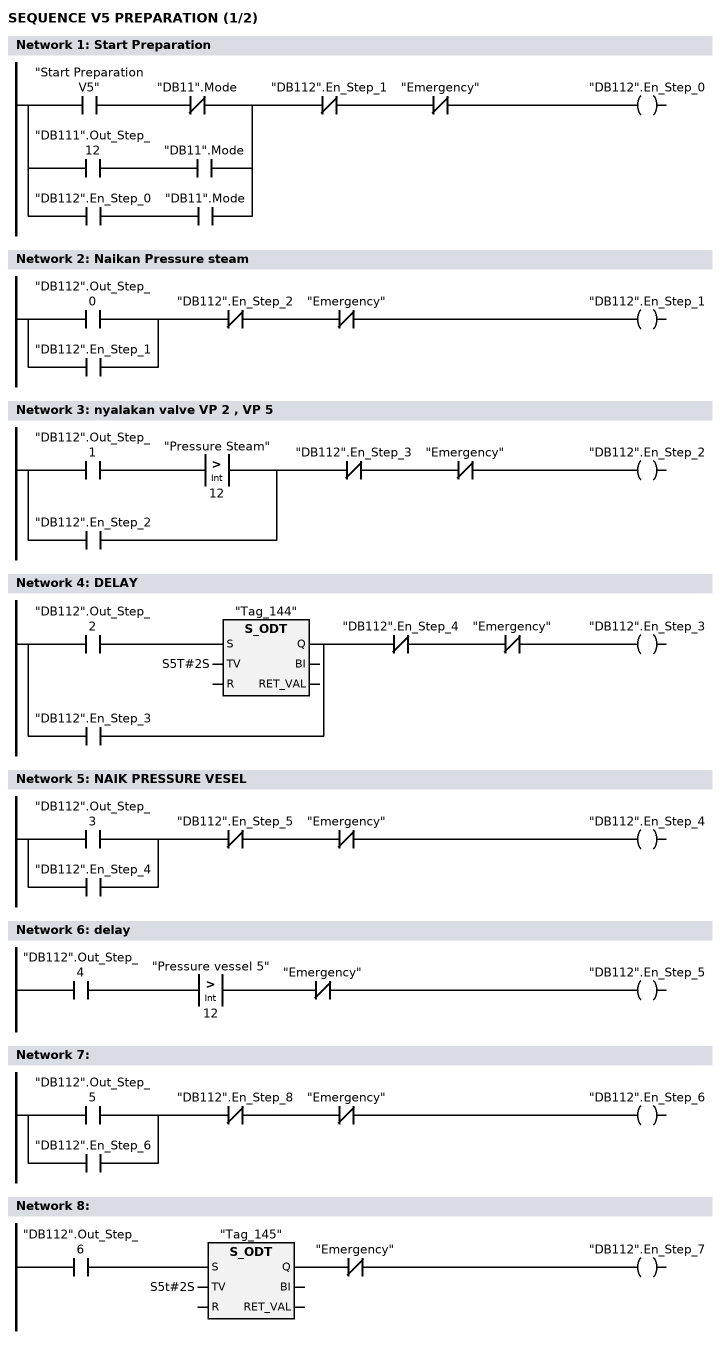
   RUNG wire#powerrail
      Contact( "Start Preparation V5" )
      I_Contact( "DB11".Mode )
      wire#w1
      I_Contact( "DB112".En_Step_1 )
      I_Contact( "Emergency" )
      Coil( "DB112".En_Step_0 )
   END_RUNG
   RUNG wire#powerrail
      Contact( "DB111".Out_Step_12 )
      Contact( "DB11".Mode )
   END_RUNG wire#w1
   RUNG wire#powerrail
      Contact( "DB112".En_Step_0 )
      Contact( "DB11".Mode )
   END_RUNG wire#w1
   // the same network as SCL:
   "DB112".En_Step_0 := (("Start Preparation V5" AND NOT "DB11".Mode) OR ("DB111".Out_Step_12 AND "DB11".Mode) OR ("DB112".En_Step_0 AND "DB11".Mode)) AND NOT "DB112".En_Step_1 AND NOT "Emergency";
END_REGION

REGION Network 2: Naikan Pressure steam
   RUNG wire#powerrail
      Contact( "DB112".Out_Step_0 )
      wire#w1
      I_Contact( "DB112".En_Step_2 )
      I_Contact( "Emergency" )
      Coil( "DB112".En_Step_1 )
   END_RUNG
   RUNG wire#powerrail
      Contact( "DB112".En_Step_1 )
   END_RUNG wire#w1
   // the same network as SCL:
   "DB112".En_Step_1 := ("DB112".Out_Step_0 OR "DB112".En_Step_1) AND NOT "DB112".En_Step_2 AND NOT "Emergency";
END_REGION

REGION Network 3: nyalakan valve VP 2 , VP 5
   RUNG wire#powerrail
      Contact( "DB112".Out_Step_1 )
      { S7_Templates := "SrcType := Int" } GT_Contact(in1 := "Pressure Steam", in2 := 12)
      wire#w1
      I_Contact( "DB112".En_Step_3 )
      I_Contact( "Emergency" )
      Coil( "DB112".En_Step_2 )
   END_RUNG
   RUNG wire#powerrail
      Contact( "DB112".En_Step_2 )
   END_RUNG wire#w1
   // the same network as SCL:
   "DB112".En_Step_2 := (("DB112".Out_Step_1 AND ("Pressure Steam" > 12)) OR "DB112".En_Step_2) AND NOT "DB112".En_Step_3 AND NOT "Emergency";
END_REGION

REGION Network 4: DELAY
   RUNG wire#powerrail
      Contact( "DB112".Out_Step_2 )
      S_ODT(T_NO := "Tag_144", TV := S5T#2S, R :=, BI =>, RET_VAL =>)
      wire#w1
      I_Contact( "DB112".En_Step_4 )
      I_Contact( "Emergency" )
      Coil( "DB112".En_Step_3 )
   END_RUNG
   RUNG wire#powerrail
      Contact( "DB112".En_Step_3 )
   END_RUNG wire#w1
   // the same network as SCL:
   #_s5time1 := S_ODT(T_NO := "Tag_144", S := "DB112".Out_Step_2, TV := S5T#2S, Q => #_w1);
   "DB112".En_Step_3 := (#_w1 OR "DB112".En_Step_3) AND NOT "DB112".En_Step_4 AND NOT "Emergency";
END_REGION

REGION Network 5: NAIK PRESSURE VESEL
   RUNG wire#powerrail
      Contact( "DB112".Out_Step_3 )
      wire#w1
      I_Contact( "DB112".En_Step_5 )
      I_Contact( "Emergency" )
      Coil( "DB112".En_Step_4 )
   END_RUNG
   RUNG wire#powerrail
      Contact( "DB112".En_Step_4 )
   END_RUNG wire#w1
   // the same network as SCL:
   "DB112".En_Step_4 := ("DB112".Out_Step_3 OR "DB112".En_Step_4) AND NOT "DB112".En_Step_5 AND NOT "Emergency";
END_REGION

REGION Network 6: delay
   RUNG wire#powerrail
      Contact( "DB112".Out_Step_4 )
      { S7_Templates := "SrcType := Int" } GT_Contact(in1 := "Pressure vessel 5", in2 := 12)
      I_Contact( "Emergency" )
      Coil( "DB112".En_Step_5 )
   END_RUNG
   // the same network as SCL:
   "DB112".En_Step_5 := "DB112".Out_Step_4 AND ("Pressure vessel 5" > 12) AND NOT "Emergency";
END_REGION

REGION Network 7
   RUNG wire#powerrail
      Contact( "DB112".Out_Step_5 )
      wire#w1
      I_Contact( "DB112".En_Step_8 )
      I_Contact( "Emergency" )
      Coil( "DB112".En_Step_6 )
   END_RUNG
   RUNG wire#powerrail
      Contact( "DB112".En_Step_6 )
   END_RUNG wire#w1
   // the same network as SCL:
   "DB112".En_Step_6 := ("DB112".Out_Step_5 OR "DB112".En_Step_6) AND NOT "DB112".En_Step_8 AND NOT "Emergency";
END_REGION

REGION Network 8
   RUNG wire#powerrail
      Contact( "DB112".Out_Step_6 )
      S_ODT(T_NO := "Tag_145", TV := S5t#2S, R :=, BI =>, RET_VAL =>)
      I_Contact( "Emergency" )
      Coil( "DB112".En_Step_7 )
   END_RUNG
   // the same network as SCL:
   #_s5time1 := S_ODT(T_NO := "Tag_145", S := "DB112".Out_Step_6, TV := S5t#2S, Q => #_w1);
   "DB112".En_Step_7 := #_w1 AND NOT "Emergency";
END_REGION

REGION Network 9: TURUNKAN PRESSURE
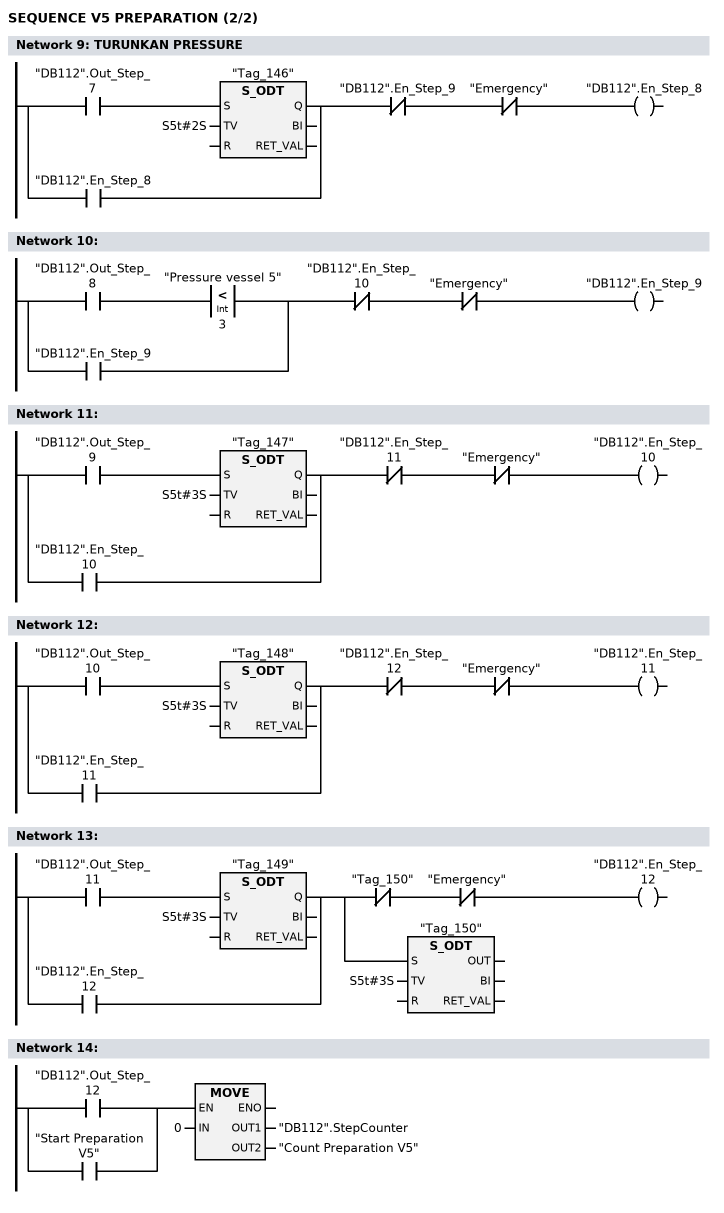
   RUNG wire#powerrail
      Contact( "DB112".Out_Step_7 )
      S_ODT(T_NO := "Tag_146", TV := S5t#2S, R :=, BI =>, RET_VAL =>)
      wire#w1
      I_Contact( "DB112".En_Step_9 )
      I_Contact( "Emergency" )
      Coil( "DB112".En_Step_8 )
   END_RUNG
   RUNG wire#powerrail
      Contact( "DB112".En_Step_8 )
   END_RUNG wire#w1
   // the same network as SCL:
   #_s5time1 := S_ODT(T_NO := "Tag_146", S := "DB112".Out_Step_7, TV := S5t#2S, Q => #_w1);
   "DB112".En_Step_8 := (#_w1 OR "DB112".En_Step_8) AND NOT "DB112".En_Step_9 AND NOT "Emergency";
END_REGION

REGION Network 10
   RUNG wire#powerrail
      Contact( "DB112".Out_Step_8 )
      { S7_Templates := "SrcType := Int" } LT_Contact(in1 := "Pressure vessel 5", in2 := 3)
      wire#w1
      I_Contact( "DB112".En_Step_10 )
      I_Contact( "Emergency" )
      Coil( "DB112".En_Step_9 )
   END_RUNG
   RUNG wire#powerrail
      Contact( "DB112".En_Step_9 )
   END_RUNG wire#w1
   // the same network as SCL:
   "DB112".En_Step_9 := (("DB112".Out_Step_8 AND ("Pressure vessel 5" < 3)) OR "DB112".En_Step_9) AND NOT "DB112".En_Step_10 AND NOT "Emergency";
END_REGION

REGION Network 11
   RUNG wire#powerrail
      Contact( "DB112".Out_Step_9 )
      S_ODT(T_NO := "Tag_147", TV := S5t#3S, R :=, BI =>, RET_VAL =>)
      wire#w1
      I_Contact( "DB112".En_Step_11 )
      I_Contact( "Emergency" )
      Coil( "DB112".En_Step_10 )
   END_RUNG
   RUNG wire#powerrail
      Contact( "DB112".En_Step_10 )
   END_RUNG wire#w1
   // the same network as SCL:
   #_s5time1 := S_ODT(T_NO := "Tag_147", S := "DB112".Out_Step_9, TV := S5t#3S, Q => #_w1);
   "DB112".En_Step_10 := (#_w1 OR "DB112".En_Step_10) AND NOT "DB112".En_Step_11 AND NOT "Emergency";
END_REGION

REGION Network 12
   RUNG wire#powerrail
      Contact( "DB112".Out_Step_10 )
      S_ODT(T_NO := "Tag_148", TV := S5t#3S, R :=, BI =>, RET_VAL =>)
      wire#w1
      I_Contact( "DB112".En_Step_12 )
      I_Contact( "Emergency" )
      Coil( "DB112".En_Step_11 )
   END_RUNG
   RUNG wire#powerrail
      Contact( "DB112".En_Step_11 )
   END_RUNG wire#w1
   // the same network as SCL:
   #_s5time1 := S_ODT(T_NO := "Tag_148", S := "DB112".Out_Step_10, TV := S5t#3S, Q => #_w1);
   "DB112".En_Step_11 := (#_w1 OR "DB112".En_Step_11) AND NOT "DB112".En_Step_12 AND NOT "Emergency";
END_REGION

REGION Network 13
   RUNG wire#powerrail
      Contact( "DB112".Out_Step_11 )
      S_ODT(T_NO := "Tag_149", TV := S5t#3S, R :=, BI =>, RET_VAL =>)
      wire#w1
      I_Contact( "Tag_150" )
      I_Contact( "Emergency" )
      Coil( "DB112".En_Step_12 )
   END_RUNG
   RUNG wire#powerrail
      Contact( "DB112".En_Step_12 )
   END_RUNG wire#w1
   RUNG wire#w1
      S_ODT(T_NO := "Tag_150", TV := S5t#3S, R :=, BI =>, RET_VAL =>)
   END_RUNG
   // the same network as SCL:
   #_s5time1 := S_ODT(T_NO := "Tag_149", S := "DB112".Out_Step_11, TV := S5t#3S, Q => #_w1);
   #_w2 := #_w1 OR "DB112".En_Step_12;
   "DB112".En_Step_12 := #_w2 AND NOT "Tag_150" AND NOT "Emergency";
   #_s5time2 := S_ODT(T_NO := "Tag_150", S := #_w2, TV := S5t#3S);
END_REGION

REGION Network 14
   RUNG wire#powerrail
      Contact( "DB112".Out_Step_12 )
      wire#w1
      Move(in := 0, out1 => "DB112".StepCounter, out2 => "Count Preparation V5")
   END_RUNG
   RUNG wire#powerrail
      Contact( "Start Preparation V5" )
   END_RUNG wire#w1
   // the same network as SCL:
   IF "DB112".Out_Step_12 OR "Start Preparation V5" THEN
       "DB112".StepCounter := 0;
       "Count Preparation V5" := 0;
   END_IF;
END_REGION
END_FUNCTION

FUNCTION "VESSEL 5 PREPARATION" : Void   // FC30, LAD
{ S7_Optimized_Access := 'TRUE' }
VERSION : 0.1
   VAR_TEMP   // added for the SCL form of the ladder/FBD networks
      _w1 : Bool;
      _w2 : Bool;
      _w3 : Bool;
      _w4 : Bool;
   END_VAR
BEGIN

REGION Network 1: NAIKAN PRESSURE STEAM
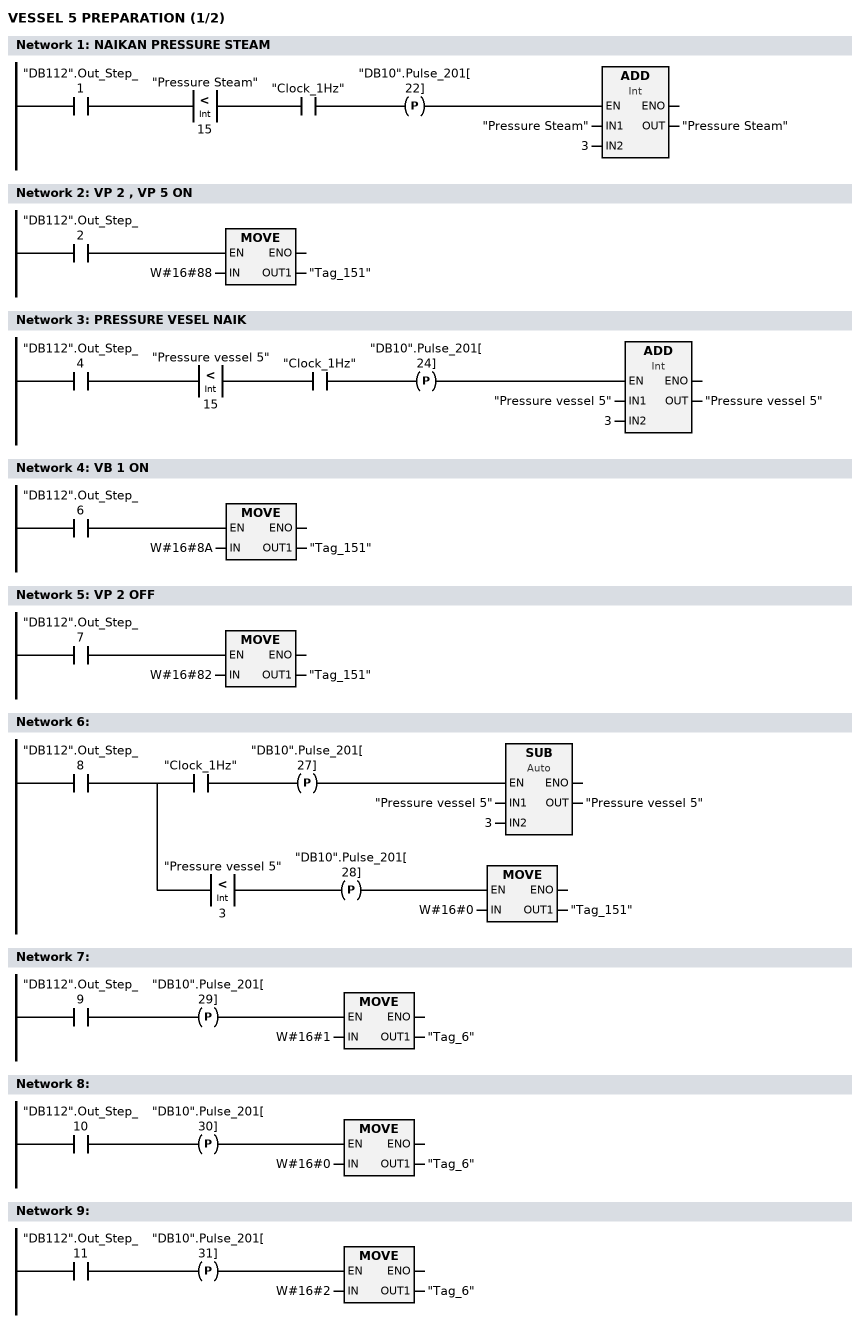
   RUNG wire#powerrail
      Contact( "DB112".Out_Step_1 )
      { S7_Templates := "SrcType := Int" } LT_Contact(in1 := "Pressure Steam", in2 := 15)
      Contact( "Clock_1Hz" )
      P_Trig( "DB10".Pulse_201[22] )
      { S7_Templates := "SrcType := Int" } Add(in1 := "Pressure Steam", in2 := 3, out => "Pressure Steam")
   END_RUNG
   // the same network as SCL:
   #_w1 := "DB112".Out_Step_1 AND ("Pressure Steam" < 15) AND "Clock_1Hz";
   #_w2 := #_w1 AND NOT "DB10".Pulse_201[22];   // rising edge
   "DB10".Pulse_201[22] := #_w1;
   IF #_w2 THEN "Pressure Steam" := "Pressure Steam" + 3; END_IF;
END_REGION

REGION Network 2: VP 2 , VP 5 ON
   RUNG wire#powerrail
      Contact( "DB112".Out_Step_2 )
      Move(in := W#16#88, out1 => "Tag_151")
   END_RUNG
   // the same network as SCL:
   IF "DB112".Out_Step_2 THEN "Tag_151" := W#16#88; END_IF;
END_REGION

REGION Network 3: PRESSURE VESEL NAIK
   RUNG wire#powerrail
      Contact( "DB112".Out_Step_4 )
      { S7_Templates := "SrcType := Int" } LT_Contact(in1 := "Pressure vessel 5", in2 := 15)
      Contact( "Clock_1Hz" )
      P_Trig( "DB10".Pulse_201[24] )
      { S7_Templates := "SrcType := Int" } Add(in1 := "Pressure vessel 5", in2 := 3, out => "Pressure vessel 5")
   END_RUNG
   // the same network as SCL:
   #_w1 := "DB112".Out_Step_4 AND ("Pressure vessel 5" < 15) AND "Clock_1Hz";
   #_w2 := #_w1 AND NOT "DB10".Pulse_201[24];   // rising edge
   "DB10".Pulse_201[24] := #_w1;
   IF #_w2 THEN "Pressure vessel 5" := "Pressure vessel 5" + 3; END_IF;
END_REGION

REGION Network 4: VB 1 ON
   RUNG wire#powerrail
      Contact( "DB112".Out_Step_6 )
      Move(in := W#16#8A, out1 => "Tag_151")
   END_RUNG
   // the same network as SCL:
   IF "DB112".Out_Step_6 THEN "Tag_151" := W#16#8A; END_IF;
END_REGION

REGION Network 5: VP 2 OFF
   RUNG wire#powerrail
      Contact( "DB112".Out_Step_7 )
      Move(in := W#16#82, out1 => "Tag_151")
   END_RUNG
   // the same network as SCL:
   IF "DB112".Out_Step_7 THEN "Tag_151" := W#16#82; END_IF;
END_REGION

REGION Network 6
   RUNG wire#powerrail
      Contact( "DB112".Out_Step_8 )
      wire#w1
      Contact( "Clock_1Hz" )
      P_Trig( "DB10".Pulse_201[27] )
      Sub(in1 := "Pressure vessel 5", in2 := 3, out => "Pressure vessel 5")
   END_RUNG
   RUNG wire#w1
      { S7_Templates := "SrcType := Int" } LT_Contact(in1 := "Pressure vessel 5", in2 := 3)
      P_Trig( "DB10".Pulse_201[28] )
      Move(in := W#16#0, out1 => "Tag_151")
   END_RUNG
   // the same network as SCL:
   #_w1 := "DB112".Out_Step_8 AND "Clock_1Hz";
   #_w2 := #_w1 AND NOT "DB10".Pulse_201[27];   // rising edge
   "DB10".Pulse_201[27] := #_w1;
   IF #_w2 THEN "Pressure vessel 5" := "Pressure vessel 5" - 3; END_IF;
   #_w3 := "DB112".Out_Step_8 AND ("Pressure vessel 5" < 3);
   #_w4 := #_w3 AND NOT "DB10".Pulse_201[28];   // rising edge
   "DB10".Pulse_201[28] := #_w3;
   IF #_w4 THEN "Tag_151" := W#16#0; END_IF;
END_REGION

REGION Network 7
   RUNG wire#powerrail
      Contact( "DB112".Out_Step_9 )
      P_Trig( "DB10".Pulse_201[29] )
      Move(in := W#16#1, out1 => "Tag_6")
   END_RUNG
   // the same network as SCL:
   #_w1 := "DB112".Out_Step_9 AND NOT "DB10".Pulse_201[29];   // rising edge
   "DB10".Pulse_201[29] := "DB112".Out_Step_9;
   IF #_w1 THEN "Tag_6" := W#16#1; END_IF;
END_REGION

REGION Network 8
   RUNG wire#powerrail
      Contact( "DB112".Out_Step_10 )
      P_Trig( "DB10".Pulse_201[30] )
      Move(in := W#16#0, out1 => "Tag_6")
   END_RUNG
   // the same network as SCL:
   #_w1 := "DB112".Out_Step_10 AND NOT "DB10".Pulse_201[30];   // rising edge
   "DB10".Pulse_201[30] := "DB112".Out_Step_10;
   IF #_w1 THEN "Tag_6" := W#16#0; END_IF;
END_REGION

REGION Network 9
   RUNG wire#powerrail
      Contact( "DB112".Out_Step_11 )
      P_Trig( "DB10".Pulse_201[31] )
      Move(in := W#16#2, out1 => "Tag_6")
   END_RUNG
   // the same network as SCL:
   #_w1 := "DB112".Out_Step_11 AND NOT "DB10".Pulse_201[31];   // rising edge
   "DB10".Pulse_201[31] := "DB112".Out_Step_11;
   IF #_w1 THEN "Tag_6" := W#16#2; END_IF;
END_REGION

REGION Network 10
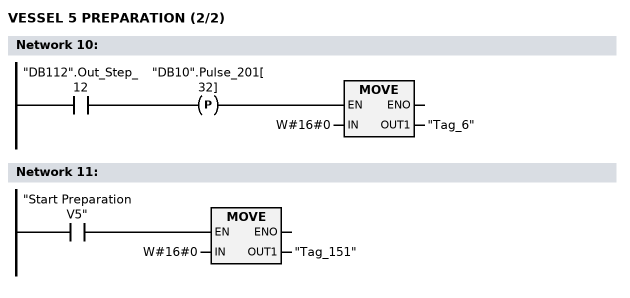
   RUNG wire#powerrail
      Contact( "DB112".Out_Step_12 )
      P_Trig( "DB10".Pulse_201[32] )
      Move(in := W#16#0, out1 => "Tag_6")
   END_RUNG
   // the same network as SCL:
   #_w1 := "DB112".Out_Step_12 AND NOT "DB10".Pulse_201[32];   // rising edge
   "DB10".Pulse_201[32] := "DB112".Out_Step_12;
   IF #_w1 THEN "Tag_6" := W#16#0; END_IF;
END_REGION

REGION Network 11
   RUNG wire#powerrail
      Contact( "Start Preparation V5" )
      Move(in := W#16#0, out1 => "Tag_151")
   END_RUNG
   // the same network as SCL:
   IF "Start Preparation V5" THEN "Tag_151" := W#16#0; END_IF;
END_REGION
END_FUNCTION

FUNCTION "SEQUENCE V6 PREPARATION" : Void   // FC31, LAD
{ S7_Optimized_Access := 'TRUE' }
VERSION : 0.1
   VAR_TEMP   // added for the SCL form of the ladder/FBD networks
      _w1 : Bool;
      _s5time1 : S5Time;
      _w2 : Bool;
      _s5time2 : S5Time;
   END_VAR
BEGIN

REGION Network 1: Start Preparation
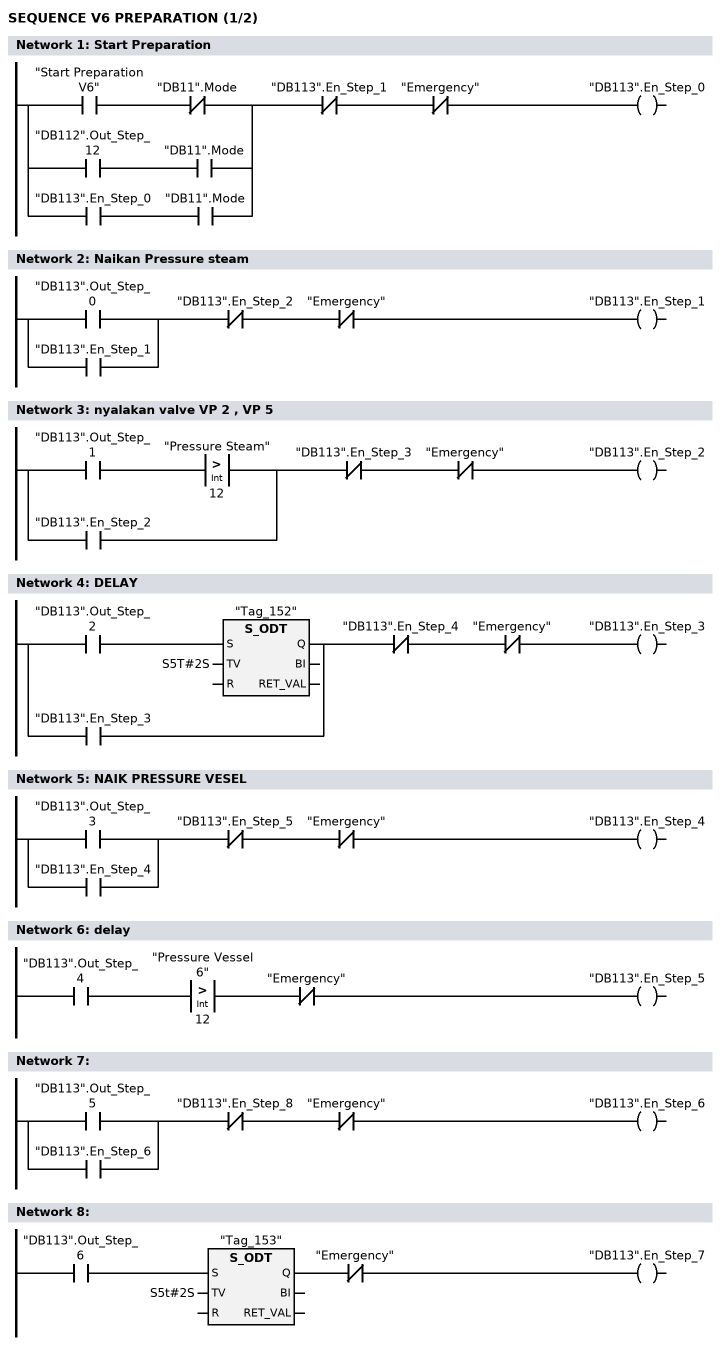
   RUNG wire#powerrail
      Contact( "Start Preparation V6" )
      I_Contact( "DB11".Mode )
      wire#w1
      I_Contact( "DB113".En_Step_1 )
      I_Contact( "Emergency" )
      Coil( "DB113".En_Step_0 )
   END_RUNG
   RUNG wire#powerrail
      Contact( "DB112".Out_Step_12 )
      Contact( "DB11".Mode )
   END_RUNG wire#w1
   RUNG wire#powerrail
      Contact( "DB113".En_Step_0 )
      Contact( "DB11".Mode )
   END_RUNG wire#w1
   // the same network as SCL:
   "DB113".En_Step_0 := (("Start Preparation V6" AND NOT "DB11".Mode) OR ("DB112".Out_Step_12 AND "DB11".Mode) OR ("DB113".En_Step_0 AND "DB11".Mode)) AND NOT "DB113".En_Step_1 AND NOT "Emergency";
END_REGION

REGION Network 2: Naikan Pressure steam
   RUNG wire#powerrail
      Contact( "DB113".Out_Step_0 )
      wire#w1
      I_Contact( "DB113".En_Step_2 )
      I_Contact( "Emergency" )
      Coil( "DB113".En_Step_1 )
   END_RUNG
   RUNG wire#powerrail
      Contact( "DB113".En_Step_1 )
   END_RUNG wire#w1
   // the same network as SCL:
   "DB113".En_Step_1 := ("DB113".Out_Step_0 OR "DB113".En_Step_1) AND NOT "DB113".En_Step_2 AND NOT "Emergency";
END_REGION

REGION Network 3: nyalakan valve VP 2 , VP 5
   RUNG wire#powerrail
      Contact( "DB113".Out_Step_1 )
      { S7_Templates := "SrcType := Int" } GT_Contact(in1 := "Pressure Steam", in2 := 12)
      wire#w1
      I_Contact( "DB113".En_Step_3 )
      I_Contact( "Emergency" )
      Coil( "DB113".En_Step_2 )
   END_RUNG
   RUNG wire#powerrail
      Contact( "DB113".En_Step_2 )
   END_RUNG wire#w1
   // the same network as SCL:
   "DB113".En_Step_2 := (("DB113".Out_Step_1 AND ("Pressure Steam" > 12)) OR "DB113".En_Step_2) AND NOT "DB113".En_Step_3 AND NOT "Emergency";
END_REGION

REGION Network 4: DELAY
   RUNG wire#powerrail
      Contact( "DB113".Out_Step_2 )
      S_ODT(T_NO := "Tag_152", TV := S5T#2S, R :=, BI =>, RET_VAL =>)
      wire#w1
      I_Contact( "DB113".En_Step_4 )
      I_Contact( "Emergency" )
      Coil( "DB113".En_Step_3 )
   END_RUNG
   RUNG wire#powerrail
      Contact( "DB113".En_Step_3 )
   END_RUNG wire#w1
   // the same network as SCL:
   #_s5time1 := S_ODT(T_NO := "Tag_152", S := "DB113".Out_Step_2, TV := S5T#2S, Q => #_w1);
   "DB113".En_Step_3 := (#_w1 OR "DB113".En_Step_3) AND NOT "DB113".En_Step_4 AND NOT "Emergency";
END_REGION

REGION Network 5: NAIK PRESSURE VESEL
   RUNG wire#powerrail
      Contact( "DB113".Out_Step_3 )
      wire#w1
      I_Contact( "DB113".En_Step_5 )
      I_Contact( "Emergency" )
      Coil( "DB113".En_Step_4 )
   END_RUNG
   RUNG wire#powerrail
      Contact( "DB113".En_Step_4 )
   END_RUNG wire#w1
   // the same network as SCL:
   "DB113".En_Step_4 := ("DB113".Out_Step_3 OR "DB113".En_Step_4) AND NOT "DB113".En_Step_5 AND NOT "Emergency";
END_REGION

REGION Network 6: delay
   RUNG wire#powerrail
      Contact( "DB113".Out_Step_4 )
      { S7_Templates := "SrcType := Int" } GT_Contact(in1 := "Pressure Vessel 6", in2 := 12)
      I_Contact( "Emergency" )
      Coil( "DB113".En_Step_5 )
   END_RUNG
   // the same network as SCL:
   "DB113".En_Step_5 := "DB113".Out_Step_4 AND ("Pressure Vessel 6" > 12) AND NOT "Emergency";
END_REGION

REGION Network 7
   RUNG wire#powerrail
      Contact( "DB113".Out_Step_5 )
      wire#w1
      I_Contact( "DB113".En_Step_8 )
      I_Contact( "Emergency" )
      Coil( "DB113".En_Step_6 )
   END_RUNG
   RUNG wire#powerrail
      Contact( "DB113".En_Step_6 )
   END_RUNG wire#w1
   // the same network as SCL:
   "DB113".En_Step_6 := ("DB113".Out_Step_5 OR "DB113".En_Step_6) AND NOT "DB113".En_Step_8 AND NOT "Emergency";
END_REGION

REGION Network 8
   RUNG wire#powerrail
      Contact( "DB113".Out_Step_6 )
      S_ODT(T_NO := "Tag_153", TV := S5t#2S, R :=, BI =>, RET_VAL =>)
      I_Contact( "Emergency" )
      Coil( "DB113".En_Step_7 )
   END_RUNG
   // the same network as SCL:
   #_s5time1 := S_ODT(T_NO := "Tag_153", S := "DB113".Out_Step_6, TV := S5t#2S, Q => #_w1);
   "DB113".En_Step_7 := #_w1 AND NOT "Emergency";
END_REGION

REGION Network 9: TURUNKAN PRESSURE
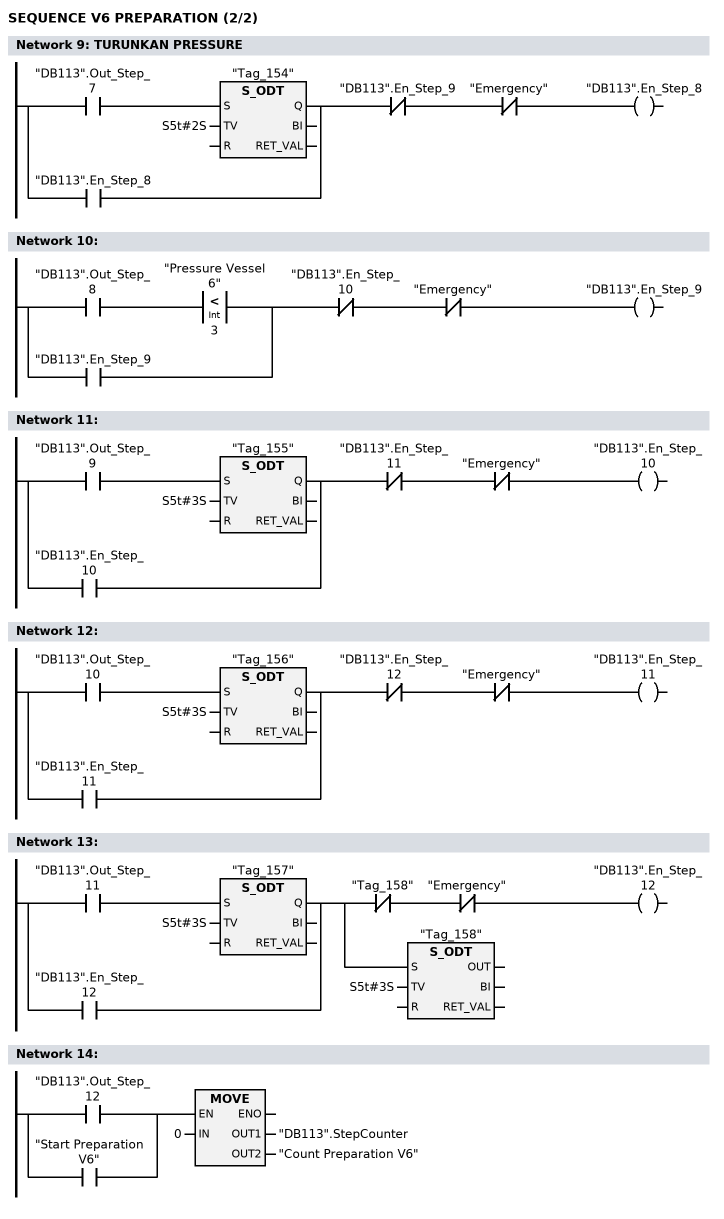
   RUNG wire#powerrail
      Contact( "DB113".Out_Step_7 )
      S_ODT(T_NO := "Tag_154", TV := S5t#2S, R :=, BI =>, RET_VAL =>)
      wire#w1
      I_Contact( "DB113".En_Step_9 )
      I_Contact( "Emergency" )
      Coil( "DB113".En_Step_8 )
   END_RUNG
   RUNG wire#powerrail
      Contact( "DB113".En_Step_8 )
   END_RUNG wire#w1
   // the same network as SCL:
   #_s5time1 := S_ODT(T_NO := "Tag_154", S := "DB113".Out_Step_7, TV := S5t#2S, Q => #_w1);
   "DB113".En_Step_8 := (#_w1 OR "DB113".En_Step_8) AND NOT "DB113".En_Step_9 AND NOT "Emergency";
END_REGION

REGION Network 10
   RUNG wire#powerrail
      Contact( "DB113".Out_Step_8 )
      { S7_Templates := "SrcType := Int" } LT_Contact(in1 := "Pressure Vessel 6", in2 := 3)
      wire#w1
      I_Contact( "DB113".En_Step_10 )
      I_Contact( "Emergency" )
      Coil( "DB113".En_Step_9 )
   END_RUNG
   RUNG wire#powerrail
      Contact( "DB113".En_Step_9 )
   END_RUNG wire#w1
   // the same network as SCL:
   "DB113".En_Step_9 := (("DB113".Out_Step_8 AND ("Pressure Vessel 6" < 3)) OR "DB113".En_Step_9) AND NOT "DB113".En_Step_10 AND NOT "Emergency";
END_REGION

REGION Network 11
   RUNG wire#powerrail
      Contact( "DB113".Out_Step_9 )
      S_ODT(T_NO := "Tag_155", TV := S5t#3S, R :=, BI =>, RET_VAL =>)
      wire#w1
      I_Contact( "DB113".En_Step_11 )
      I_Contact( "Emergency" )
      Coil( "DB113".En_Step_10 )
   END_RUNG
   RUNG wire#powerrail
      Contact( "DB113".En_Step_10 )
   END_RUNG wire#w1
   // the same network as SCL:
   #_s5time1 := S_ODT(T_NO := "Tag_155", S := "DB113".Out_Step_9, TV := S5t#3S, Q => #_w1);
   "DB113".En_Step_10 := (#_w1 OR "DB113".En_Step_10) AND NOT "DB113".En_Step_11 AND NOT "Emergency";
END_REGION

REGION Network 12
   RUNG wire#powerrail
      Contact( "DB113".Out_Step_10 )
      S_ODT(T_NO := "Tag_156", TV := S5t#3S, R :=, BI =>, RET_VAL =>)
      wire#w1
      I_Contact( "DB113".En_Step_12 )
      I_Contact( "Emergency" )
      Coil( "DB113".En_Step_11 )
   END_RUNG
   RUNG wire#powerrail
      Contact( "DB113".En_Step_11 )
   END_RUNG wire#w1
   // the same network as SCL:
   #_s5time1 := S_ODT(T_NO := "Tag_156", S := "DB113".Out_Step_10, TV := S5t#3S, Q => #_w1);
   "DB113".En_Step_11 := (#_w1 OR "DB113".En_Step_11) AND NOT "DB113".En_Step_12 AND NOT "Emergency";
END_REGION

REGION Network 13
   RUNG wire#powerrail
      Contact( "DB113".Out_Step_11 )
      S_ODT(T_NO := "Tag_157", TV := S5t#3S, R :=, BI =>, RET_VAL =>)
      wire#w1
      I_Contact( "Tag_158" )
      I_Contact( "Emergency" )
      Coil( "DB113".En_Step_12 )
   END_RUNG
   RUNG wire#powerrail
      Contact( "DB113".En_Step_12 )
   END_RUNG wire#w1
   RUNG wire#w1
      S_ODT(T_NO := "Tag_158", TV := S5t#3S, R :=, BI =>, RET_VAL =>)
   END_RUNG
   // the same network as SCL:
   #_s5time1 := S_ODT(T_NO := "Tag_157", S := "DB113".Out_Step_11, TV := S5t#3S, Q => #_w1);
   #_w2 := #_w1 OR "DB113".En_Step_12;
   "DB113".En_Step_12 := #_w2 AND NOT "Tag_158" AND NOT "Emergency";
   #_s5time2 := S_ODT(T_NO := "Tag_158", S := #_w2, TV := S5t#3S);
END_REGION

REGION Network 14
   RUNG wire#powerrail
      Contact( "DB113".Out_Step_12 )
      wire#w1
      Move(in := 0, out1 => "DB113".StepCounter, out2 => "Count Preparation V6")
   END_RUNG
   RUNG wire#powerrail
      Contact( "Start Preparation V6" )
   END_RUNG wire#w1
   // the same network as SCL:
   IF "DB113".Out_Step_12 OR "Start Preparation V6" THEN
       "DB113".StepCounter := 0;
       "Count Preparation V6" := 0;
   END_IF;
END_REGION
END_FUNCTION

FUNCTION "VESSEL 6 PREPARATION" : Void   // FC32, LAD
{ S7_Optimized_Access := 'TRUE' }
VERSION : 0.1
   VAR_TEMP   // added for the SCL form of the ladder/FBD networks
      _w1 : Bool;
      _w2 : Bool;
      _w3 : Bool;
      _w4 : Bool;
   END_VAR
BEGIN

REGION Network 1: NAIKAN PRESSURE STEAM
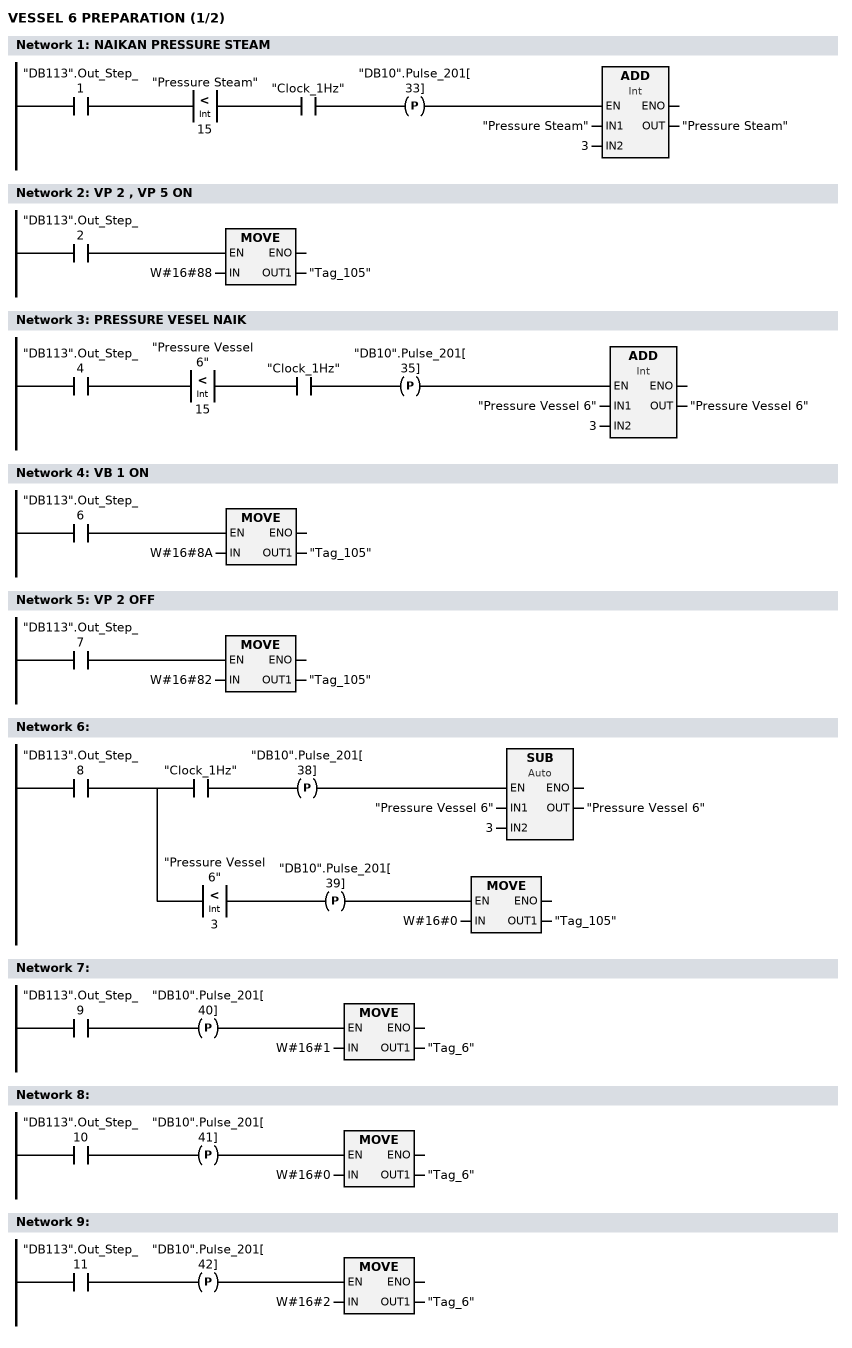
   RUNG wire#powerrail
      Contact( "DB113".Out_Step_1 )
      { S7_Templates := "SrcType := Int" } LT_Contact(in1 := "Pressure Steam", in2 := 15)
      Contact( "Clock_1Hz" )
      P_Trig( "DB10".Pulse_201[33] )
      { S7_Templates := "SrcType := Int" } Add(in1 := "Pressure Steam", in2 := 3, out => "Pressure Steam")
   END_RUNG
   // the same network as SCL:
   #_w1 := "DB113".Out_Step_1 AND ("Pressure Steam" < 15) AND "Clock_1Hz";
   #_w2 := #_w1 AND NOT "DB10".Pulse_201[33];   // rising edge
   "DB10".Pulse_201[33] := #_w1;
   IF #_w2 THEN "Pressure Steam" := "Pressure Steam" + 3; END_IF;
END_REGION

REGION Network 2: VP 2 , VP 5 ON
   RUNG wire#powerrail
      Contact( "DB113".Out_Step_2 )
      Move(in := W#16#88, out1 => "Tag_105")
   END_RUNG
   // the same network as SCL:
   IF "DB113".Out_Step_2 THEN "Tag_105" := W#16#88; END_IF;
END_REGION

REGION Network 3: PRESSURE VESEL NAIK
   RUNG wire#powerrail
      Contact( "DB113".Out_Step_4 )
      { S7_Templates := "SrcType := Int" } LT_Contact(in1 := "Pressure Vessel 6", in2 := 15)
      Contact( "Clock_1Hz" )
      P_Trig( "DB10".Pulse_201[35] )
      { S7_Templates := "SrcType := Int" } Add(in1 := "Pressure Vessel 6", in2 := 3, out => "Pressure Vessel 6")
   END_RUNG
   // the same network as SCL:
   #_w1 := "DB113".Out_Step_4 AND ("Pressure Vessel 6" < 15) AND "Clock_1Hz";
   #_w2 := #_w1 AND NOT "DB10".Pulse_201[35];   // rising edge
   "DB10".Pulse_201[35] := #_w1;
   IF #_w2 THEN "Pressure Vessel 6" := "Pressure Vessel 6" + 3; END_IF;
END_REGION

REGION Network 4: VB 1 ON
   RUNG wire#powerrail
      Contact( "DB113".Out_Step_6 )
      Move(in := W#16#8A, out1 => "Tag_105")
   END_RUNG
   // the same network as SCL:
   IF "DB113".Out_Step_6 THEN "Tag_105" := W#16#8A; END_IF;
END_REGION

REGION Network 5: VP 2 OFF
   RUNG wire#powerrail
      Contact( "DB113".Out_Step_7 )
      Move(in := W#16#82, out1 => "Tag_105")
   END_RUNG
   // the same network as SCL:
   IF "DB113".Out_Step_7 THEN "Tag_105" := W#16#82; END_IF;
END_REGION

REGION Network 6
   RUNG wire#powerrail
      Contact( "DB113".Out_Step_8 )
      wire#w1
      Contact( "Clock_1Hz" )
      P_Trig( "DB10".Pulse_201[38] )
      Sub(in1 := "Pressure Vessel 6", in2 := 3, out => "Pressure Vessel 6")
   END_RUNG
   RUNG wire#w1
      { S7_Templates := "SrcType := Int" } LT_Contact(in1 := "Pressure Vessel 6", in2 := 3)
      P_Trig( "DB10".Pulse_201[39] )
      Move(in := W#16#0, out1 => "Tag_105")
   END_RUNG
   // the same network as SCL:
   #_w1 := "DB113".Out_Step_8 AND "Clock_1Hz";
   #_w2 := #_w1 AND NOT "DB10".Pulse_201[38];   // rising edge
   "DB10".Pulse_201[38] := #_w1;
   IF #_w2 THEN "Pressure Vessel 6" := "Pressure Vessel 6" - 3; END_IF;
   #_w3 := "DB113".Out_Step_8 AND ("Pressure Vessel 6" < 3);
   #_w4 := #_w3 AND NOT "DB10".Pulse_201[39];   // rising edge
   "DB10".Pulse_201[39] := #_w3;
   IF #_w4 THEN "Tag_105" := W#16#0; END_IF;
END_REGION

REGION Network 7
   RUNG wire#powerrail
      Contact( "DB113".Out_Step_9 )
      P_Trig( "DB10".Pulse_201[40] )
      Move(in := W#16#1, out1 => "Tag_6")
   END_RUNG
   // the same network as SCL:
   #_w1 := "DB113".Out_Step_9 AND NOT "DB10".Pulse_201[40];   // rising edge
   "DB10".Pulse_201[40] := "DB113".Out_Step_9;
   IF #_w1 THEN "Tag_6" := W#16#1; END_IF;
END_REGION

REGION Network 8
   RUNG wire#powerrail
      Contact( "DB113".Out_Step_10 )
      P_Trig( "DB10".Pulse_201[41] )
      Move(in := W#16#0, out1 => "Tag_6")
   END_RUNG
   // the same network as SCL:
   #_w1 := "DB113".Out_Step_10 AND NOT "DB10".Pulse_201[41];   // rising edge
   "DB10".Pulse_201[41] := "DB113".Out_Step_10;
   IF #_w1 THEN "Tag_6" := W#16#0; END_IF;
END_REGION

REGION Network 9
   RUNG wire#powerrail
      Contact( "DB113".Out_Step_11 )
      P_Trig( "DB10".Pulse_201[42] )
      Move(in := W#16#2, out1 => "Tag_6")
   END_RUNG
   // the same network as SCL:
   #_w1 := "DB113".Out_Step_11 AND NOT "DB10".Pulse_201[42];   // rising edge
   "DB10".Pulse_201[42] := "DB113".Out_Step_11;
   IF #_w1 THEN "Tag_6" := W#16#2; END_IF;
END_REGION

REGION Network 10